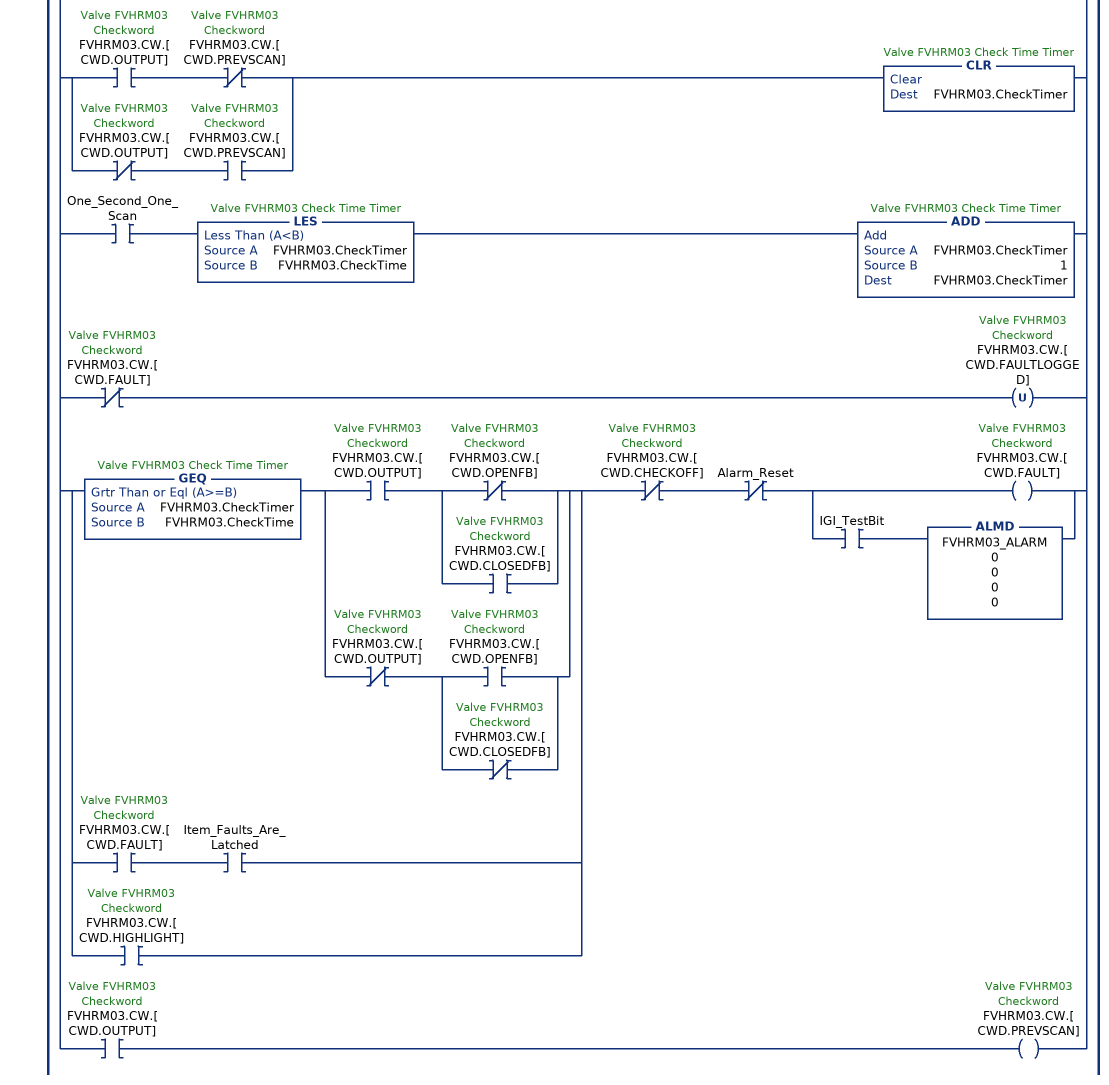
   85: [NEQ(FVHRM03.DriveBits,0) OTE(FVHRM03.CW.[CWD.AUTODRV]) ,[XIC(FVHRM03.CW.[CWD.AUTODRV]) XIO(FVHRM03.CW.[CWD.MANUAL]) ,XIC(FVHRM03.CW.[CWD.MANDRV]) XIC(FVHRM03.CW.[CWD.MANUAL]) ] OTE(FVHRM03.CW.[CWD.OUTPUT]) ,XIC(FVHRM03.CW.[CWD.OUTPUT]) OTE(FVHRM03_DR) ,XIC(S:FS) [OTU(FVHRM03.CW.[CWD.MANUAL]) ,LEQ(FVHRM03.CheckTime,0) MOV(Default_Check_Time,FVHRM03.CheckTime) ] ,[[XIC(FVHRM03_OP) XIO(Item_Simulation_Flag) ,XIC(Item_Simulation_Flag) XIC(FVHRM03.CW.[CWD.OUTPUT]) XIO(FVHRM03.CW.[CWD.SIMFAIL]) ] OTE(FVHRM03.CW.[CWD.OPENFB]) ,[XIC(FVHRM03_CL) XIO(Item_Simulation_Flag) ,XIC(Item_Simulation_Flag) XIO(FVHRM03.CW.[CWD.OUTPUT]) XIO(FVHRM03.CW.[CWD.SIMFAIL]) ] OTE(FVHRM03.CW.[CWD.CLOSEDFB]) ] ,[XIC(FVHRM03.CW.[CWD.OUTPUT]) XIO(FVHRM03.CW.[CWD.PREVSCAN]) ,XIO(FVHRM03.CW.[CWD.OUTPUT]) XIC(FVHRM03.CW.[CWD.PREVSCAN]) ] CLR(FVHRM03.CheckTimer) ,XIC(One_Second_One_Scan) LES(FVHRM03.CheckTimer,FVHRM03.CheckTime) ADD(FVHRM03.CheckTimer,1,FVHRM03.CheckTimer) ,XIO(FVHRM03.CW.[CWD.FAULT]) OTU(FVHRM03.CW.[CWD.FAULTLOGGED]) ,[GEQ(FVHRM03.CheckTimer,FVHRM03.CheckTime) [XIC(FVHRM03.CW.[CWD.OUTPUT]) [XIO(FVHRM03.CW.[CWD.OPENFB]) ,XIC(FVHRM03.CW.[CWD.CLOSEDFB]) ] ,XIO(FVHRM03.CW.[CWD.OUTPUT]) [XIC(FVHRM03.CW.[CWD.OPENFB]) ,XIO(FVHRM03.CW.[CWD.CLOSEDFB]) ] ] ,XIC(FVHRM03.CW.[CWD.FAULT]) XIC(Item_Faults_Are_Latched) ,XIC(FVHRM03.CW.[CWD.HIGHLIGHT]) ] XIO(FVHRM03.CW.[CWD.CHECKOFF]) XIO(Alarm_Reset) [OTE(FVHRM03.CW.[CWD.FAULT]) ,XIC(IGI_TestBit) ALMD(FVHRM03_ALARM,0,0,0,0) ] ,XIC(FVHRM03.CW.[CWD.OUTPUT]) OTE(FVHRM03.CW.[CWD.PREVSCAN]) ];
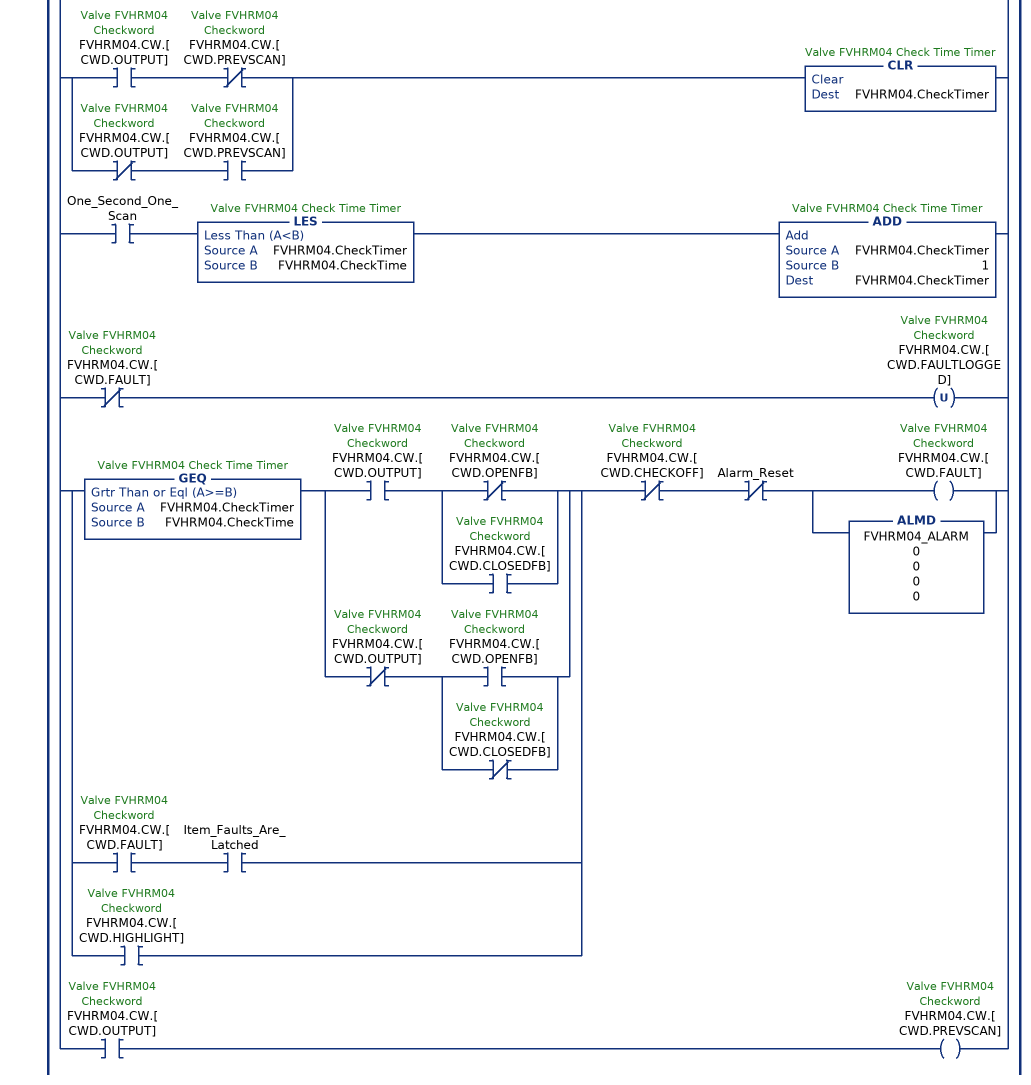
   86: [NEQ(FVHRM04.DriveBits,0) OTE(FVHRM04.CW.[CWD.AUTODRV]) ,[XIC(FVHRM04.CW.[CWD.AUTODRV]) XIO(FVHRM04.CW.[CWD.MANUAL]) ,XIC(FVHRM04.CW.[CWD.MANDRV]) XIC(FVHRM04.CW.[CWD.MANUAL]) ] OTE(FVHRM04.CW.[CWD.OUTPUT]) ,XIC(FVHRM04.CW.[CWD.OUTPUT]) OTE(FVHRM04_DR) ,XIC(S:FS) [OTU(FVHRM04.CW.[CWD.MANUAL]) ,LEQ(FVHRM04.CheckTime,0) MOV(Default_Check_Time,FVHRM04.CheckTime) ] ,[[XIC(FVHRM04_OP) XIO(Item_Simulation_Flag) ,XIC(Item_Simulation_Flag) XIC(FVHRM04.CW.[CWD.OUTPUT]) XIO(FVHRM04.CW.[CWD.SIMFAIL]) ] OTE(FVHRM04.CW.[CWD.OPENFB]) ,[XIC(FVHRM04_CL) XIO(Item_Simulation_Flag) ,XIC(Item_Simulation_Flag) XIO(FVHRM04.CW.[CWD.OUTPUT]) XIO(FVHRM04.CW.[CWD.SIMFAIL]) ] OTE(FVHRM04.CW.[CWD.CLOSEDFB]) ] ,[XIC(FVHRM04.CW.[CWD.OUTPUT]) XIO(FVHRM04.CW.[CWD.PREVSCAN]) ,XIO(FVHRM04.CW.[CWD.OUTPUT]) XIC(FVHRM04.CW.[CWD.PREVSCAN]) ] CLR(FVHRM04.CheckTimer) ,XIC(One_Second_One_Scan) LES(FVHRM04.CheckTimer,FVHRM04.CheckTime) ADD(FVHRM04.CheckTimer,1,FVHRM04.CheckTimer) ,XIO(FVHRM04.CW.[CWD.FAULT]) OTU(FVHRM04.CW.[CWD.FAULTLOGGED]) ,[GEQ(FVHRM04.CheckTimer,FVHRM04.CheckTime) [XIC(FVHRM04.CW.[CWD.OUTPUT]) [XIO(FVHRM04.CW.[CWD.OPENFB]) ,XIC(FVHRM04.CW.[CWD.CLOSEDFB]) ] ,XIO(FVHRM04.CW.[CWD.OUTPUT]) [XIC(FVHRM04.CW.[CWD.OPENFB]) ,XIO(FVHRM04.CW.[CWD.CLOSEDFB]) ] ] ,XIC(FVHRM04.CW.[CWD.FAULT]) XIC(Item_Faults_Are_Latched) ,XIC(FVHRM04.CW.[CWD.HIGHLIGHT]) ] XIO(FVHRM04.CW.[CWD.CHECKOFF]) XIO(Alarm_Reset) [OTE(FVHRM04.CW.[CWD.FAULT]) ,ALMD(FVHRM04_ALARM,0,0,0,0) ] ,XIC(FVHRM04.CW.[CWD.OUTPUT]) OTE(FVHRM04.CW.[CWD.PREVSCAN]) ];
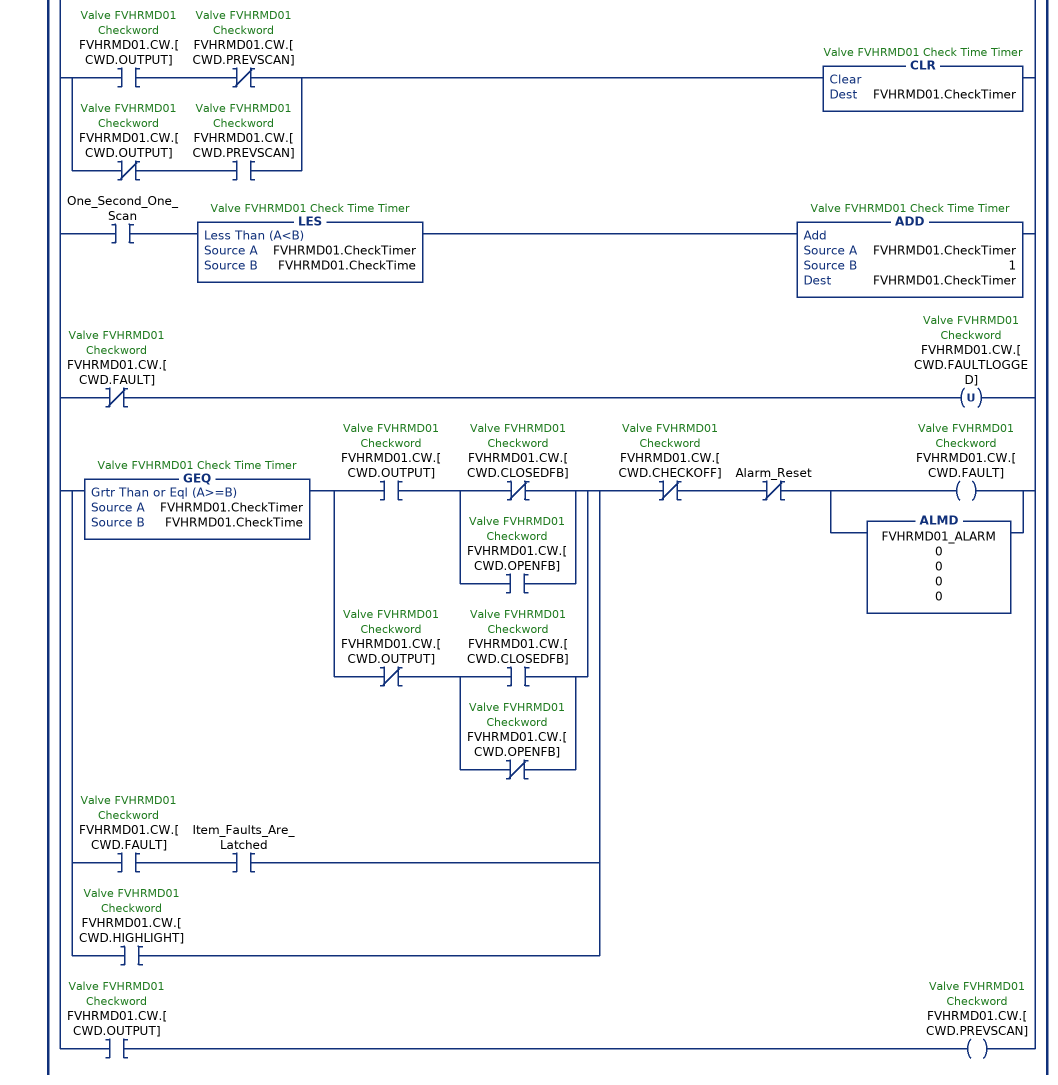
   87: [NEQ(FVHRMD01.DriveBits,0) OTE(FVHRMD01.CW.[CWD.AUTODRV]) ,[XIC(FVHRMD01.CW.[CWD.AUTODRV]) XIO(FVHRMD01.CW.[CWD.MANUAL]) ,XIC(FVHRMD01.CW.[CWD.MANDRV]) XIC(FVHRMD01.CW.[CWD.MANUAL]) ] OTE(FVHRMD01.CW.[CWD.OUTPUT]) ,XIC(FVHRMD01.CW.[CWD.OUTPUT]) OTE(FVHRMD01_DR) ,XIC(S:FS) [OTU(FVHRMD01.CW.[CWD.MANUAL]) ,LEQ(FVHRMD01.CheckTime,0) MOV(Default_Check_Time,FVHRMD01.CheckTime) ] ,[[XIC(FVHRMD01_OP) XIO(Item_Simulation_Flag) ,XIC(Item_Simulation_Flag) XIC(FVHRMD01.CW.[CWD.OUTPUT]) XIO(FVHRMD01.CW.[CWD.SIMFAIL]) ] OTE(FVHRMD01.CW.[CWD.OPENFB]) ,[XIC(FVHRMD01_CL) XIO(Item_Simulation_Flag) ,XIC(Item_Simulation_Flag) XIO(FVHRMD01.CW.[CWD.OUTPUT]) XIO(FVHRMD01.CW.[CWD.SIMFAIL]) ] OTE(FVHRMD01.CW.[CWD.CLOSEDFB]) ] ,[XIC(FVHRMD01.CW.[CWD.OUTPUT]) XIO(FVHRMD01.CW.[CWD.PREVSCAN]) ,XIO(FVHRMD01.CW.[CWD.OUTPUT]) XIC(FVHRMD01.CW.[CWD.PREVSCAN]) ] CLR(FVHRMD01.CheckTimer) ,XIC(One_Second_One_Scan) LES(FVHRMD01.CheckTimer,FVHRMD01.CheckTime) ADD(FVHRMD01.CheckTimer,1,FVHRMD01.CheckTimer) ,XIO(FVHRMD01.CW.[CWD.FAULT]) OTU(FVHRMD01.CW.[CWD.FAULTLOGGED]) ,[GEQ(FVHRMD01.CheckTimer,FVHRMD01.CheckTime) [XIC(FVHRMD01.CW.[CWD.OUTPUT]) [XIO(FVHRMD01.CW.[CWD.CLOSEDFB]) ,XIC(FVHRMD01.CW.[CWD.OPENFB]) ] ,XIO(FVHRMD01.CW.[CWD.OUTPUT]) [XIC(FVHRMD01.CW.[CWD.CLOSEDFB]) ,XIO(FVHRMD01.CW.[CWD.OPENFB]) ] ] ,XIC(FVHRMD01.CW.[CWD.FAULT]) XIC(Item_Faults_Are_Latched) ,XIC(FVHRMD01.CW.[CWD.HIGHLIGHT]) ] XIO(FVHRMD01.CW.[CWD.CHECKOFF]) XIO(Alarm_Reset) [OTE(FVHRMD01.CW.[CWD.FAULT]) ,ALMD(FVHRMD01_ALARM,0,0,0,0) ] ,XIC(FVHRMD01.CW.[CWD.OUTPUT]) OTE(FVHRMD01.CW.[CWD.PREVSCAN]) ];
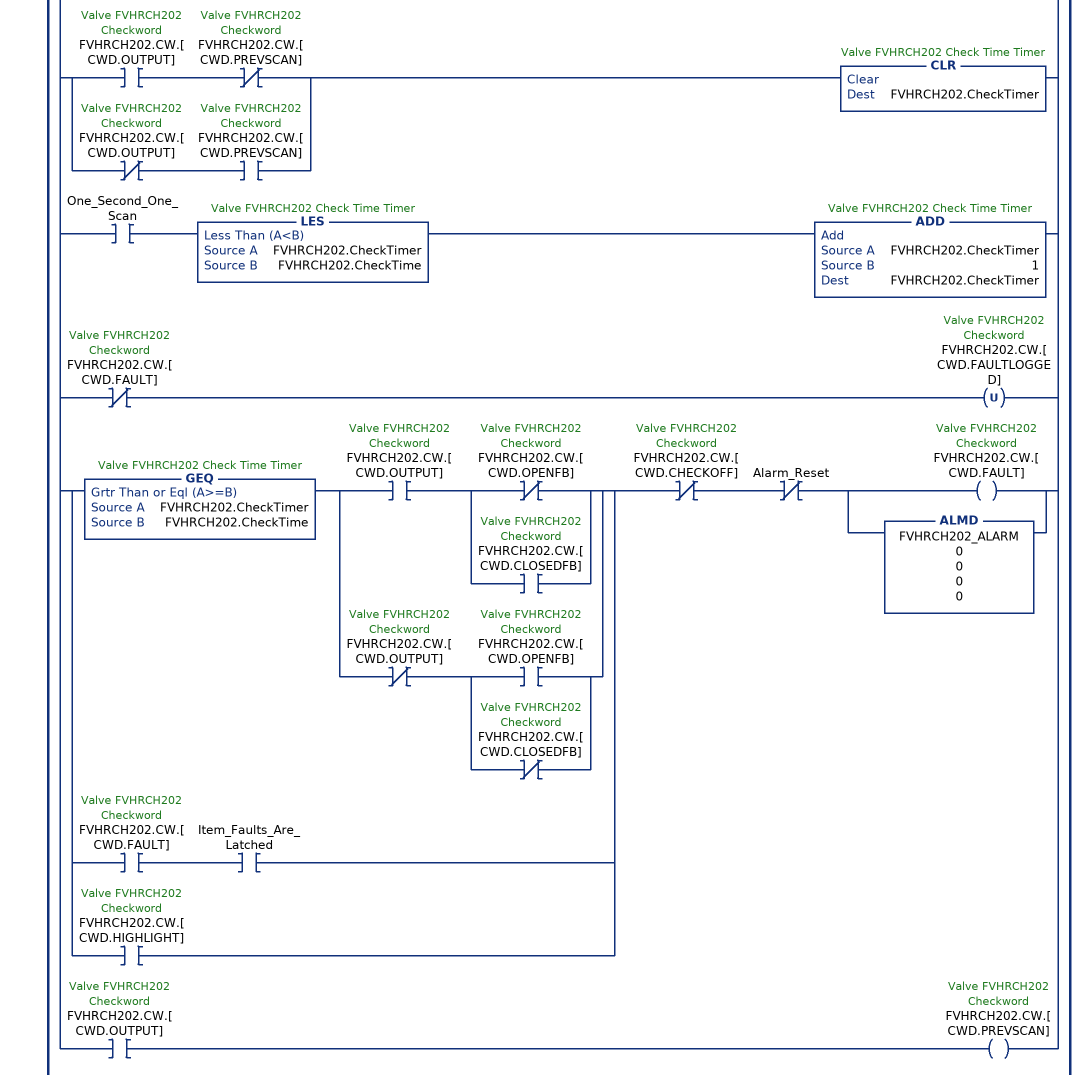
   88: [NEQ(FVHRCH202.DriveBits,0) OTE(FVHRCH202.CW.[CWD.AUTODRV]) ,[XIC(FVHRCH202.CW.[CWD.AUTODRV]) XIO(FVHRCH202.CW.[CWD.MANUAL]) ,XIC(FVHRCH202.CW.[CWD.MANDRV]) XIC(FVHRCH202.CW.[CWD.MANUAL]) ] OTE(FVHRCH202.CW.[CWD.OUTPUT]) ,XIC(FVHRCH202.CW.[CWD.OUTPUT]) OTE(FVHRCH202_DR) ,XIC(S:FS) [OTU(FVHRCH202.CW.[CWD.MANUAL]) ,LEQ(FVHRCH202.CheckTime,0) MOV(Default_Check_Time,FVHRCH202.CheckTime) ] ,[[XIC(FVHRCH202_OP) XIO(Item_Simulation_Flag) ,XIC(Item_Simulation_Flag) XIC(FVHRCH202.CW.[CWD.OUTPUT]) XIO(FVHRCH202.CW.[CWD.SIMFAIL]) ] OTE(FVHRCH202.CW.[CWD.OPENFB]) ,[XIC(FVHRCH202_CL) XIO(Item_Simulation_Flag) ,XIC(Item_Simulation_Flag) XIO(FVHRCH202.CW.[CWD.OUTPUT]) XIO(FVHRCH202.CW.[CWD.SIMFAIL]) ] OTE(FVHRCH202.CW.[CWD.CLOSEDFB]) ] ,[XIC(FVHRCH202.CW.[CWD.OUTPUT]) XIO(FVHRCH202.CW.[CWD.PREVSCAN]) ,XIO(FVHRCH202.CW.[CWD.OUTPUT]) XIC(FVHRCH202.CW.[CWD.PREVSCAN]) ] CLR(FVHRCH202.CheckTimer) ,XIC(One_Second_One_Scan) LES(FVHRCH202.CheckTimer,FVHRCH202.CheckTime) ADD(FVHRCH202.CheckTimer,1,FVHRCH202.CheckTimer) ,XIO(FVHRCH202.CW.[CWD.FAULT]) OTU(FVHRCH202.CW.[CWD.FAULTLOGGED]) ,[GEQ(FVHRCH202.CheckTimer,FVHRCH202.CheckTime) [XIC(FVHRCH202.CW.[CWD.OUTPUT]) [XIO(FVHRCH202.CW.[CWD.OPENFB]) ,XIC(FVHRCH202.CW.[CWD.CLOSEDFB]) ] ,XIO(FVHRCH202.CW.[CWD.OUTPUT]) [XIC(FVHRCH202.CW.[CWD.OPENFB]) ,XIO(FVHRCH202.CW.[CWD.CLOSEDFB]) ] ] ,XIC(FVHRCH202.CW.[CWD.FAULT]) XIC(Item_Faults_Are_Latched) ,XIC(FVHRCH202.CW.[CWD.HIGHLIGHT]) ] XIO(FVHRCH202.CW.[CWD.CHECKOFF]) XIO(Alarm_Reset) [OTE(FVHRCH202.CW.[CWD.FAULT]) ,ALMD(FVHRCH202_ALARM,0,0,0,0) ] ,XIC(FVHRCH202.CW.[CWD.OUTPUT]) OTE(FVHRCH202.CW.[CWD.PREVSCAN]) ];
END_ROUTINE
END_PROGRAM

PROGRAM MV_Common   (* main routine MainRoutine *)

ROUTINE A_SecondsToHMS   (* ladder *)
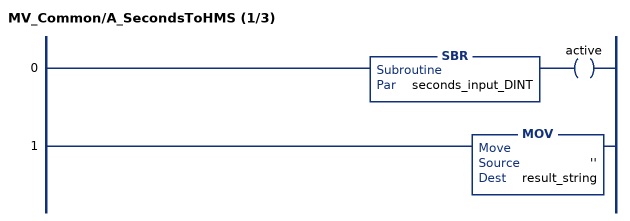
   0: SBR(seconds_input_DINT)OTE(active);
   1: MOV('',result_string);
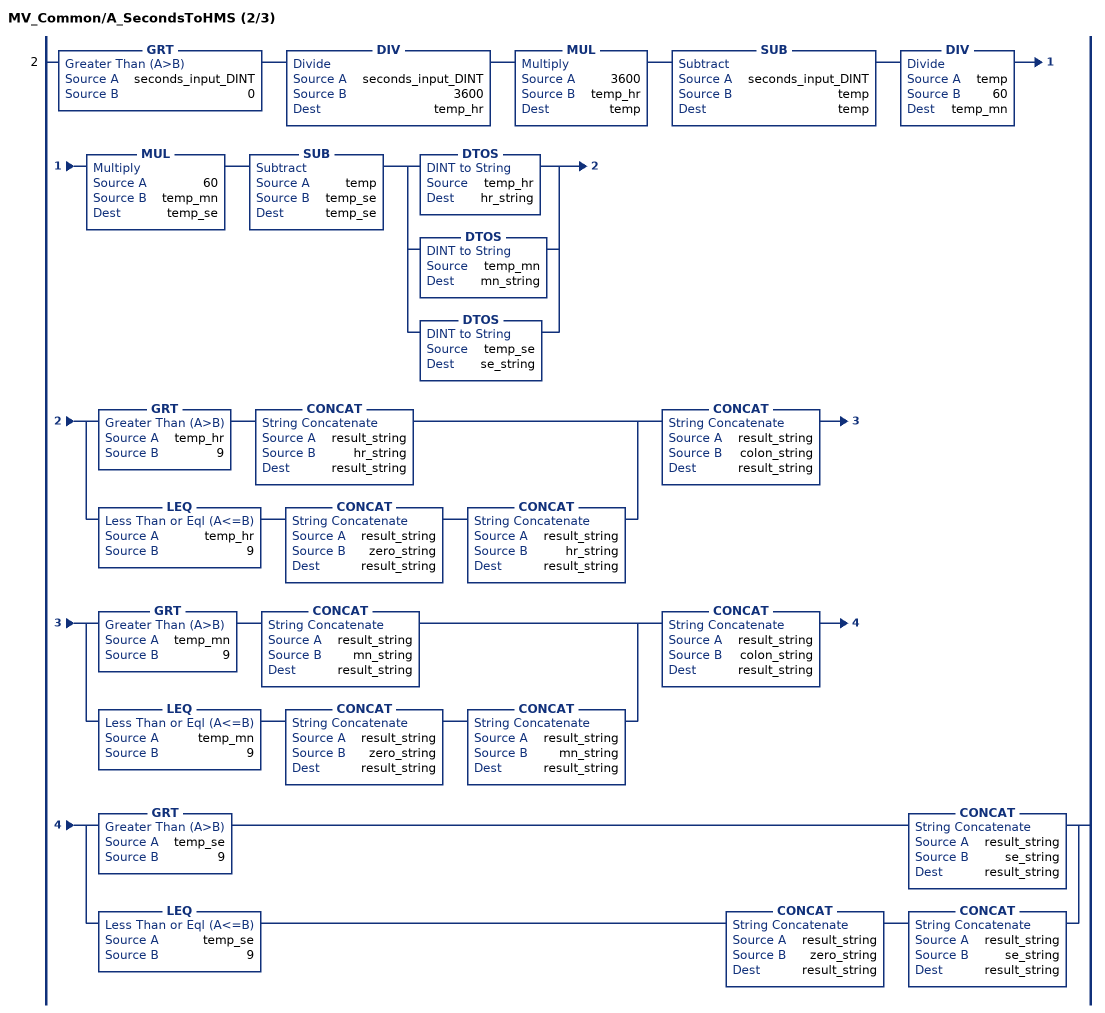
   2: GRT(seconds_input_DINT,0)DIV(seconds_input_DINT,3600,temp_hr)MUL(3600,temp_hr,temp)SUB(seconds_input_DINT,temp,temp)DIV(temp,60,temp_mn)MUL(60,temp_mn,temp_se)SUB(temp,temp_se,temp_se)[DTOS(temp_hr,hr_string) ,DTOS(temp_mn,mn_string) ,DTOS(temp_se,se_string) ][GRT(temp_hr,9) CONCAT(result_string,hr_string,result_string) ,LEQ(temp_hr,9) CONCAT(result_string,zero_string,result_string) CONCAT(result_string,hr_string,result_string) ]CONCAT(result_string,colon_string,result_string)[GRT(temp_mn,9) CONCAT(result_string,mn_string,result_string) ,LEQ(temp_mn,9) CONCAT(result_string,zero_string,result_string) CONCAT(result_string,mn_string,result_string) ]CONCAT(result_string,colon_string,result_string)[GRT(temp_se,9) CONCAT(result_string,se_string,result_string) ,LEQ(temp_se,9) CONCAT(result_string,zero_string,result_string) CONCAT(result_string,se_string,result_string) ];
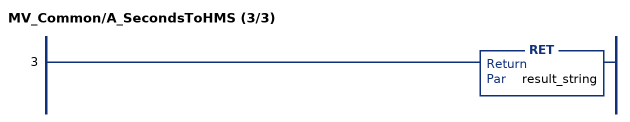
   3: RET(result_string);
END_ROUTINE

ROUTINE Analog_scale_ftof   (* ladder *)
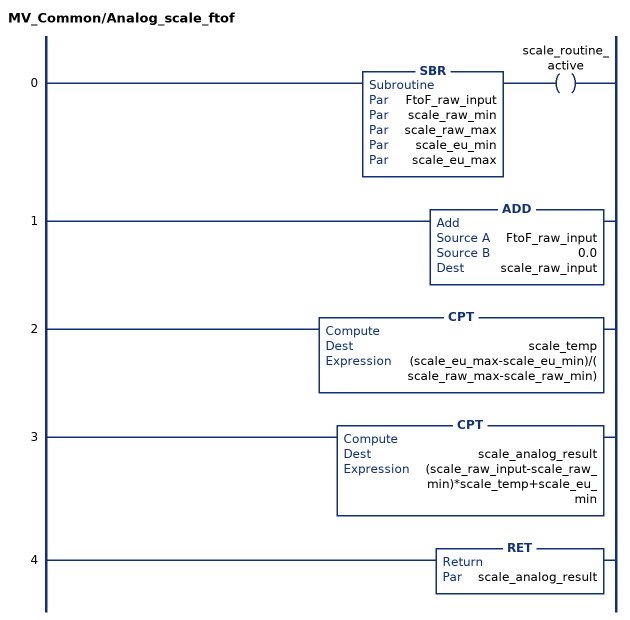
   0: SBR(FtoF_raw_input,scale_raw_min,scale_raw_max,scale_eu_min,scale_eu_max)OTE(scale_routine_active);
   1: ADD(FtoF_raw_input,0.0,scale_raw_input);
   2: CPT(scale_temp,(scale_eu_max-scale_eu_min)/(scale_raw_max-scale_raw_min));
   3: CPT(scale_analog_result,(scale_raw_input-scale_raw_min)*scale_temp+scale_eu_min);
   4: RET(scale_analog_result);
END_ROUTINE

ROUTINE Analog_Scale_FtoI   (* ladder *)
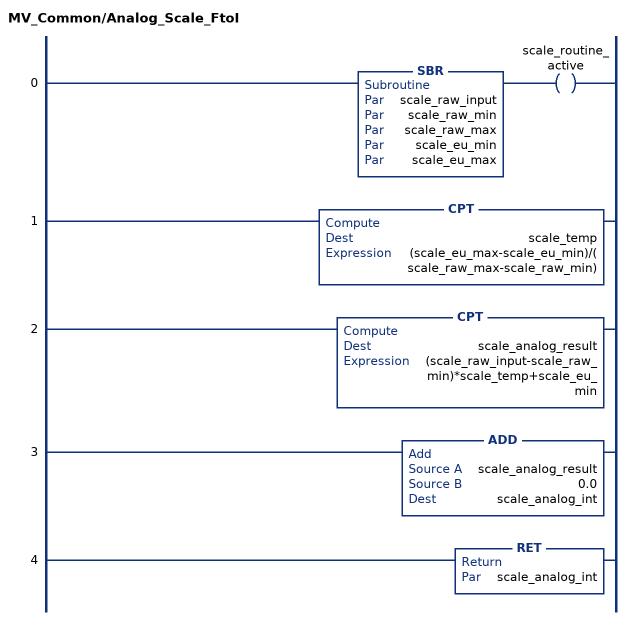
   0: SBR(scale_raw_input,scale_raw_min,scale_raw_max,scale_eu_min,scale_eu_max)OTE(scale_routine_active);
   1: CPT(scale_temp,(scale_eu_max-scale_eu_min)/(scale_raw_max-scale_raw_min));
   2: CPT(scale_analog_result,(scale_raw_input-scale_raw_min)*scale_temp+scale_eu_min);
   3: ADD(scale_analog_result,0.0,scale_analog_int);
   4: RET(scale_analog_int);
END_ROUTINE

ROUTINE Analog_Scale_ItoF   (* ladder *)
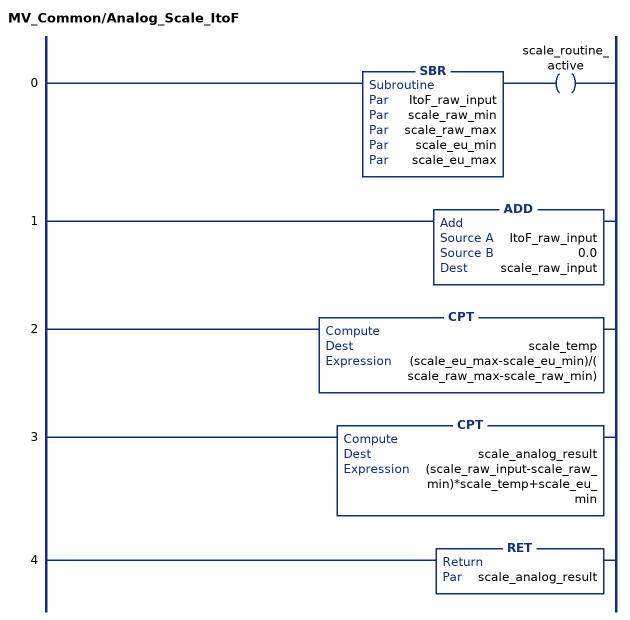
   0: SBR(ItoF_raw_input,scale_raw_min,scale_raw_max,scale_eu_min,scale_eu_max)OTE(scale_routine_active);
   1: ADD(ItoF_raw_input,0.0,scale_raw_input);
   2: CPT(scale_temp,(scale_eu_max-scale_eu_min)/(scale_raw_max-scale_raw_min));
   3: CPT(scale_analog_result,(scale_raw_input-scale_raw_min)*scale_temp+scale_eu_min);
   4: RET(scale_analog_result);
END_ROUTINE

ROUTINE ClockRoutines   (* ladder *)
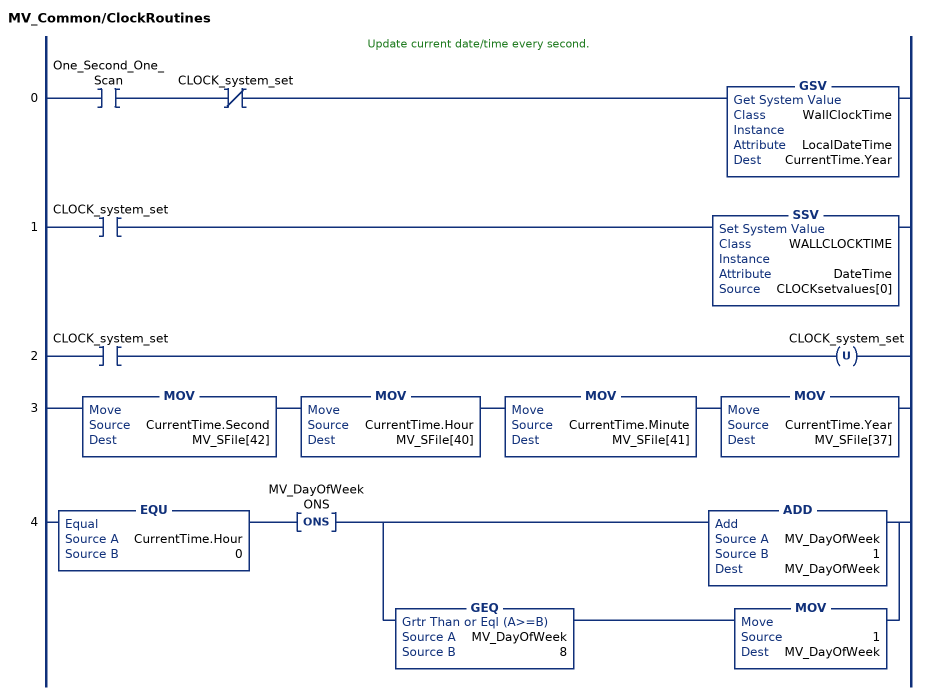
   // Update current date/time every second.
   0: XIC(One_Second_One_Scan)XIO(CLOCK_system_set)GSV(WallClockTime,,LocalDateTime,CurrentTime.Year);
   1: XIC(CLOCK_system_set)SSV(WALLCLOCKTIME,,DateTime,CLOCKsetvalues[0]);
   2: XIC(CLOCK_system_set)OTU(CLOCK_system_set);
   3: MOV(CurrentTime.Second,MV_SFile[42])MOV(CurrentTime.Hour,MV_SFile[40])MOV(CurrentTime.Minute,MV_SFile[41])MOV(CurrentTime.Year,MV_SFile[37]);
   4: EQU(CurrentTime.Hour,0)ONS(MV_DayOfWeekONS)[ADD(MV_DayOfWeek,1,MV_DayOfWeek) ,GEQ(MV_DayOfWeek,8) MOV(1,MV_DayOfWeek) ];
END_ROUTINE

ROUTINE Constants   (* ladder *)
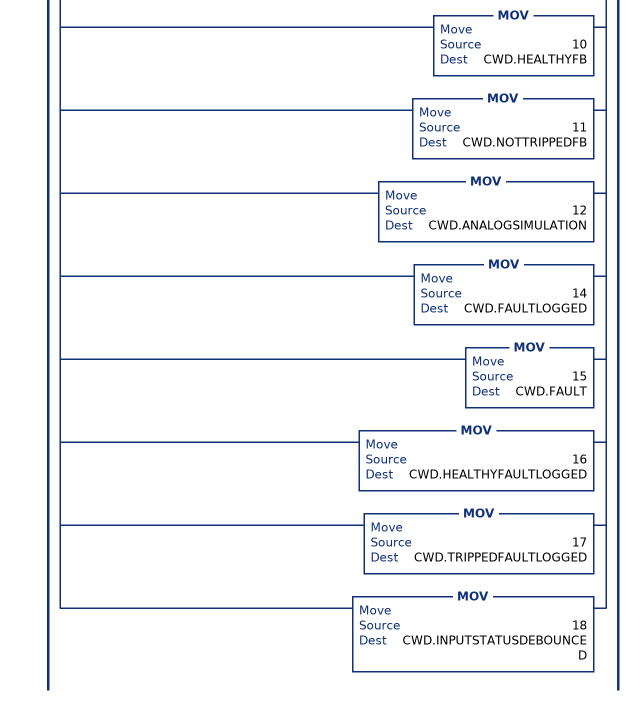
   0: [MOV(0,CWD.AUTODRV) ,MOV(0,CWD.INPUTSTATUS) ,MOV(1,CWD.PREVSCAN) ,MOV(2,CWD.SIMFAIL) ,MOV(3,CWD.OPENFB) ,MOV(3,CWD.RUNFB) ,MOV(4,CWD.CLOSEDFB) ,MOV(5,CWD.MANDRV) ,MOV(6,CWD.MANUAL) ,MOV(7,CWD.OUTPUT) ,MOV(8,CWD.CHECKOFF) ,MOV(9,CWD.HIGHLIGHT) ,MOV(10,CWD.HEALTHYFB) ,MOV(11,CWD.NOTTRIPPEDFB) ,MOV(12,CWD.ANALOGSIMULATION) ,MOV(14,CWD.FAULTLOGGED) ,MOV(15,CWD.FAULT) ,MOV(16,CWD.HEALTHYFAULTLOGGED) ,MOV(17,CWD.TRIPPEDFAULTLOGGED) ,MOV(18,CWD.INPUTSTATUSDEBOUNCED) ];
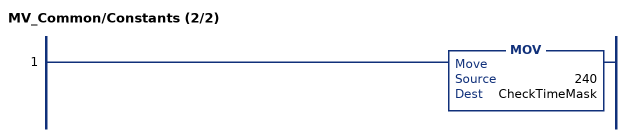
   1: MOV(240,CheckTimeMask);
END_ROUTINE
